
   REGION OUTPUTS
     // Write outputs
     IF (#statDisablingCompleted = TRUE) THEN
       // Reset outputs if disabling completed
       #statValid := FALSE;
       #statBusy := FALSE;
       #statError := FALSE;
       #statErrorUserCleared := FALSE;
       #statErrorAutoCleared := FALSE;
       #statStatus := #STATUS_NO_CALL;
       // TODO: Reset application specific outputs
       #statWaitMain := FALSE;

     ELSIF (#statErrorUserCleared = TRUE) AND (#statError = FALSE) THEN
       // Error can only be cleared by user; rising edge at enable input is needed to continue 
       #statValid := FALSE;
       #statBusy := FALSE;
       #statError := TRUE;
       #statFBState := #FB_STATE_NO_PROCESSING; // Switch state machine to "no processing"

     ELSIF (#statErrorAutoCleared = TRUE) AND (#statError = FALSE) THEN
       // Error can be reset by FB automatically  
       #statValid := FALSE;
       #statBusy := TRUE;
       #statError := TRUE;
       // TODO: Handling of autocleared error

     ELSIF (#statErrorAutoCleared = FALSE) AND (#statErrorUserCleared = FALSE) AND (#statError = TRUE) THEN
       // If autocleared error is acknowledged
       #statValid := TRUE;
       #statBusy := TRUE;
       #statError := FALSE;
       #statStatus := #STATUS_SUBSEQUENT_CALL;
     END_IF;

     // Write static values to outputs
     #valid := #statValid;
     #busy := #statBusy;
     #error := #statError;
     #status := #statStatus;
     // TODO: Write application specific static values to outputs
     #waitMain := #statWaitMain;
   END_REGION OUTPUTS
END_FUNCTION_BLOCK

FUNCTION "LKinCtrl_CheckPathDataCmd" : Word   // FC35000, SCL
TITLE = LKinCtrl_CheckPathDataCmd
{ S7_Optimized_Access := 'TRUE' }
AUTHOR : tech.team.motioncontrol@siemens.com
FAMILY : LKinCtrl
VERSION : 1.3
// The FC checks a PathData command to be configured correctly
   VAR_OUTPUT
      cmdIsMotionCmd : Bool;   // TRUE: Command is a motion command
   END_VAR
   VAR_IN_OUT
      pathDataCmd : Variant;   // variant for PathData command
   END_VAR
   VAR_TEMP
      tmpError : Bool;   // temporary variable for error bit
      tmpStatus : Word;   // temporary variable for status word
      tempFlagCtr : Int;   // temporary counter for flags
      tempPathDataCmd_regular : REF_TO "LKinCtrl_typePathDataElement";   // temporary reference to PathData element
      tempPathDataCmd_PreBuf : REF_TO "LKinCtrl_typePathDataElement_PreBuf";   // temporary reference to PathData_PreBuf element
      tempPathDataCmd_checking : "LKinCtrl_typePathDataElement";   // temporary variable for PathDataElement being checked
      tempPathDataType : Int;   // temporary variable storing detected PathData type
   END_VAR
   // Ret_Val : return value
   VAR CONSTANT
      STATUS_NO_ERROR_IN_COMMAND : Word := 16#0000;   // status no error found command
      ERR_PATHDATA_CMDTYPE : Word := 16#80A0;   // error due to wrong cmdType
      ERR_PATHDATA_COORDSYSTEM : Word := 16#80B1;   // error due to wrong coordinate system
      ERR_PATHDATA_VELOCITY : Word := 16#8003;   // error due to wrong velocity
      ERR_PATHDATA_ACCELERATION : Word := 16#8004;   // error due to wrong acceleration
      ERR_PATHDATA_DECELERATION : Word := 16#8005;   // error due to wrong deceleration
      ERR_PATHDATA_JERK : Word := 16#8006;   // error due to wrong jerk
      ERR_PATHDATA_ORIENTATIONDIRECTION : Word := 16#8007;   // error due to wrong orientation direction
      ERR_PATHDATA_BUFFERMODE : Word := 16#80B2;   // error due to wrong buffer mode
      ERR_PATHDATA_DYNAMICADAPTION : Word := 16#80B5;   // error due to wrong dynamic adaption
      ERR_PATHDATA_CIRCMODE : Word := 16#80B6;   // error due to wrong circle mode
      ERR_PATHDATA_PATHCHOICE : Word := 16#80B9;   // error due to wrong path choice
      ERR_PATHDATA_CIRCLEPLANE : Word := 16#80BA;   // error due to wrong circle plane
      ERR_PATHDATA_RADIUS : Word := 16#80BB;   // error due to wrong radius
      ERR_PATHDATA_ARC : Word := 16#80BC;   // error due to wrong arc
      ERR_PATHDATA_SETFLAGS_FLAG : Word := 16#80D1;   // error due to wrong set flag definition
      ERR_PATHDATA_SETFLAGS_FLAGMODE : Word := 16#80D2;   // error due to wrong set flag mode definition
      ERR_PATHDATA_VALUEFLAGS_FLAG : Word := 16#80D3;   // error due to wrong value flag definition
      ERR_PATHDATA_VALUEFLAGS_FLAGMODE : Word := 16#80D4;   // error due to wrong value flag mode definition
      ERR_PATHDATA_OFFSET_PARA_NO : Word := 16#80A1;   // error due to wrong offset parameter set number
      ERR_PATHDATA_OFFSET_MAINPATHPLANE : Word := 16#80A2;   // error due to wrong main path plane
      ERR_PATHDATA_POSITIONMODE : Word := 16#80A3;   // error due to wrong position mode
      ERR_PATHDATA_LINK_CONSTELLATION : Word := 16#80A4;   // error due to wrong link constellation
      ERR_PATHDATA_CONVEYOR_PARA_NO : Word := 16#80A5;   // error due to wrong conveyor parameter set number / error due to wrong link constellation
   END_VAR
BEGIN
   //==========================================================================================
   // SIEMENS AG
   // (c)Copyright 2020 All Rights Reserved
   //------------------------------------------------------------------------------------------
   // Library: LKinCtrl
   // Tested with: S7-1517T-3 PN/DP
   // Engineering: TIA Portal V15
   // Restrictions: ---
   // Requirements: S7-1500T FW 2.8
   // Functionality: LKinCtrl_CheckPathDataCmd
   // The FC checks a PathData command to be configured correctly
   // 
   // Support: tech.team.motioncontrol@siemens.com
   // Note: Parameter comments are only available in language 'English (United States)'
   //------------------------------------------------------------------------------------------
   // Change log table:
   // Version    Date          Expert in charge    Changes applied
   // 01.00.00   26.02.2019    JR                  First release version v1.0
   // 01.01.00   14.06.2019    JR                  added flagOnly command
   // 01.02.00   03.12.2019    JR                  added command checks for value flags
   // 01.02.01   30.01.2020    FR                  separate constant for flag arrays
   // 01.02.02   09.04.2020    FR                  copy valueFlags & CS to temp also
   // 01.03.00   16.04.2020    FR                  added moveDirect & trackConveyor
   //===========================================================================================

   // FC initialization
   //====================================================================================================================================
   #tmpError := FALSE;
   #tmpStatus := #STATUS_NO_ERROR_IN_COMMAND;

   // PathData conversion (reduced, regular(no suffix), advanced)
   //===========================================================================================
   REGION PATHDATA_ELEMENT_CONVERSION
     // regulat PathDataCommand
       IF TypeOf(#pathDataCmd) = LKinCtrl_typePathDataElement THEN
           // reference internal PathDataCommand to attached Variant
           #tempPathDataCmd_regular ?= #pathDataCmd;
           #tempPathDataType := 1;
           // copy to internal PathData (full version)
           #tempPathDataCmd_checking.cmdType := #tempPathDataCmd_regular<?OpDeref?>.cmdType;
           #tempPathDataCmd_checking.cmdCoordinates.coordSystem := #tempPathDataCmd_regular<?OpDeref?>.cmdCoordinates.coordSystem;
           #tempPathDataCmd_checking.cmdParameters := #tempPathDataCmd_regular<?OpDeref?>.cmdParameters;
           #tempPathDataCmd_checking.setFlags := #tempPathDataCmd_regular<?OpDeref?>.setFlags;
           #tempPathDataCmd_checking.valueFlags := #tempPathDataCmd_regular<?OpDeref?>.valueFlags;

           // PathDataPreBuffered PathDataCommand
       ELSIF TypeOf(#pathDataCmd) = LKinCtrl_typePathDataElement_PreBuf THEN
           #tempPathDataCmd_PreBuf ?= #pathDataCmd;
           #tempPathDataType := 2;
           // copy to internal PathData (full version)
           #tempPathDataCmd_checking.cmdType := #tempPathDataCmd_PreBuf<?OpDeref?>.cmdType;
           #tempPathDataCmd_checking.cmdCoordinates.coordSystem := #tempPathDataCmd_PreBuf<?OpDeref?>.cmdCoordinates.coordSystem;
           #tempPathDataCmd_checking.cmdParameters := #tempPathDataCmd_PreBuf<?OpDeref?>.cmdParameters;
           #tempPathDataCmd_checking.setFlags := #tempPathDataCmd_PreBuf<?OpDeref?>.setFlags;
           #tempPathDataCmd_checking.valueFlags := #tempPathDataCmd_PreBuf<?OpDeref?>.valueFlags;
       END_IF;
   END_REGION PATHDATA_CONVERSION 

   // PathData command 
   //====================================================================================================================================
   //PathData - command - cmdType
   // check for wrong PathData parameter cmdType
   IF (#tempPathDataCmd_checking.cmdType < "LKINCTRL_CMD_FLAG_ONLY"                      // lower limit MC cmdTypes
       OR #tempPathDataCmd_checking.cmdType > "LKINCTRL_MC_MOVEDIRECTREL")               // upper limit MC cmdTypes
     AND #tempPathDataCmd_checking.cmdType <> "LKINCTRL_CMD_WAIT_TIME"                   // exact cmdType constant for wait time
     AND #tempPathDataCmd_checking.cmdType <> "LKINCTRL_CONFIG_START_OFFSET_COMP_LEFT"   // exact cmdType constant for activation offset compensation left
     AND #tempPathDataCmd_checking.cmdType <> "LKINCTRL_CONFIG_START_OFFSET_COMP_RIGHT"  // exact cmdType constant for activation offset compensation right
     AND #tempPathDataCmd_checking.cmdType <> "LKINCTRL_CONFIG_END_OFFSET_COMP"          // exact cmdType constant for deactivation offset compensation
     AND #tempPathDataCmd_checking.cmdType <> "LKINCTRL_MC_TRACKCONVEYORBELT"
   THEN
     #tmpError := TRUE;
     #tmpStatus := #ERR_PATHDATA_CMDTYPE;
   END_IF;

   //PathData - command - cmdType
   // add separation for motion / non-motion commands here
   IF #tempPathDataCmd_checking.cmdType = "LKINCTRL_CMD_WAIT_TIME"
       OR #tempPathDataCmd_checking.cmdType = "LKINCTRL_CMD_FLAG_ONLY"
       OR #tempPathDataCmd_checking.cmdType = "LKINCTRL_MC_TRACKCONVEYORBELT"
     // add further non-motion commands here later (Zones, CS, ...)
     // only separate commands that will be copied to PathData_preBuffered
   THEN
     #cmdIsMotionCmd := FALSE;
   ELSE
     #cmdIsMotionCmd := TRUE;
   END_IF;

   //PathData - command - cmdCoordinates - coordSystem
   IF #tempPathDataCmd_checking.cmdType >= "LKINCTRL_MC_MOVELINEARABS"                           // lower limit path command cmdTypes
       AND #tempPathDataCmd_checking.cmdType <= "LKINCTRL_MC_MOVECIRCULARREL"                    // upper limit path command cmdTypes
   THEN
       // check for wrong parameter PathData coordSystem
       // CS is not WCS - OCS3 --> Error
       IF #tempPathDataCmd_checking.cmdCoordinates.coordSystem < "CS_WCS"
           OR #tempPathDataCmd_checking.cmdCoordinates.coordSystem > "CS_OCS3"
       THEN
           #tmpError := TRUE;
           #tmpStatus := #ERR_PATHDATA_COORDSYSTEM;
       END_IF;
   ELSIF #tempPathDataCmd_checking.cmdType >= "LKINCTRL_MC_MOVEDIRECTABS"                          // lower limit axis command cmdTypes
       AND #tempPathDataCmd_checking.cmdType <= "LKINCTRL_MC_MOVEDIRECTREL"                        // upper limit axis command cmdTypes
   THEN
       // check for wrong parameter PathData coordSystem
       // CS is not WCS - OCS3 and not MCS --> Error
       IF (#tempPathDataCmd_checking.cmdCoordinates.coordSystem < "CS_WCS"
           OR #tempPathDataCmd_checking.cmdCoordinates.coordSystem > "CS_OCS3")
           AND NOT (#tempPathDataCmd_checking.cmdCoordinates.coordSystem = "CS_MCS")
       THEN
           #tmpError := TRUE;
           #tmpStatus := #ERR_PATHDATA_COORDSYSTEM;
       END_IF;
       // Check conveyTracking coordinate system to be OCS1-3
   ELSIF #tempPathDataCmd_checking.cmdType = "LKINCTRL_MC_TRACKCONVEYORBELT"
       AND (#tempPathDataCmd_checking.cmdCoordinates.coordSystem < "CS_OCS1"
       OR #tempPathDataCmd_checking.cmdCoordinates.coordSystem > "CS_OCS3")
   THEN
       #tmpError := TRUE;
       #tmpStatus := #ERR_PATHDATA_COORDSYSTEM;
   END_IF;

   //PathData - command - cmdParameters - pathDynamics
   // Check MoveDirect dynamics
   IF #tempPathDataCmd_checking.cmdType >= "LKINCTRL_MC_MOVEDIRECTABS"                          // lower limit axis command cmdTypes
       AND #tempPathDataCmd_checking.cmdType <= "LKINCTRL_MC_MOVEDIRECTREL"                     // upper limit axis command cmdTypes
   THEN                
       // Check for wrong dynamics factors
       IF #tempPathDataCmd_checking.cmdParameters.pathDynamics.velocity > 1.0
           OR #tempPathDataCmd_checking.cmdParameters.pathDynamics.velocity = 0.0
       THEN
           #tmpError := TRUE;
           #tmpStatus := #ERR_PATHDATA_VELOCITY;
       END_IF;
       IF #tempPathDataCmd_checking.cmdParameters.pathDynamics.acceleration > 1.0
           OR #tempPathDataCmd_checking.cmdParameters.pathDynamics.acceleration = 0.0
       THEN
           #tmpError := TRUE;
           #tmpStatus := #ERR_PATHDATA_ACCELERATION;
       END_IF;
       IF #tempPathDataCmd_checking.cmdParameters.pathDynamics.deceleration > 1.0
           OR #tempPathDataCmd_checking.cmdParameters.pathDynamics.deceleration = 0.0
       THEN
           #tmpError := TRUE;
           #tmpStatus := #ERR_PATHDATA_DECELERATION;
       END_IF;
       IF (#tempPathDataCmd_checking.cmdParameters.pathDynamics.jerk > 0.0
           AND #tempPathDataCmd_checking.cmdParameters.pathDynamics.jerk < 0.1)
           OR #tempPathDataCmd_checking.cmdParameters.pathDynamics.jerk > 0.9
       THEN
           #tmpError := TRUE;
           #tmpStatus := #ERR_PATHDATA_JERK;
       END_IF;
   END_IF;

   //PathData - command - cmdParameters - orientationDirection
   // check for wrong parameter PathData orientationDirection
   IF #tempPathDataCmd_checking.cmdParameters.orientationDirection < 1
     OR #tempPathDataCmd_checking.cmdParameters.orientationDirection > 3
   THEN
     #tmpError := TRUE;
     #tmpStatus := #ERR_PATHDATA_ORIENTATIONDIRECTION;
   END_IF;

   //PathData - command - cmdParameters - bufferMode
   // check for wrong parameter PathData bufferMode
   IF #tempPathDataCmd_checking.cmdParameters.bufferMode <> 1
     AND #tempPathDataCmd_checking.cmdParameters.bufferMode <> 2
     AND #tempPathDataCmd_checking.cmdParameters.bufferMode <> 5
   THEN
     #tmpError := TRUE;
     #tmpStatus := #ERR_PATHDATA_BUFFERMODE;
   END_IF;

   //PathData - command - cmdParameters - dynamicAdaption
   // check for wrong parameter PathData dynamicAdaption
   IF #tempPathDataCmd_checking.cmdParameters.dynamicAdaption > 2
   THEN
     #tmpError := TRUE;
     #tmpStatus := #ERR_PATHDATA_DYNAMICADAPTION;
   END_IF;

   //PathData - command - circleParameter
   //====================================================================================================================================
   //PathData - command - circleParameter - circMode
   // check for wrong parameter PathData circMode
   IF #tempPathDataCmd_checking.cmdParameters.circleParameters.circMode < 0
     OR #tempPathDataCmd_checking.cmdParameters.circleParameters.circMode > 3
   THEN
     #tmpError := TRUE;
     #tmpStatus := #ERR_PATHDATA_CIRCMODE;
   END_IF;

   //PathData - command - circleParameter - pathChoice
   // check for wrong parameter PathData pathChoice
   IF #tempPathDataCmd_checking.cmdParameters.circleParameters.pathChoice < 0
     OR #tempPathDataCmd_checking.cmdParameters.circleParameters.pathChoice > 3
   THEN
     #tmpError := TRUE;
     #tmpStatus := #ERR_PATHDATA_PATHCHOICE;
   END_IF;

   //PathData - command - circleParameter - circlePlane
   // check for wrong parameter PathData circlePlane
   IF #tempPathDataCmd_checking.cmdParameters.circleParameters.circlePlane < 0
     OR #tempPathDataCmd_checking.cmdParameters.circleParameters.circlePlane > 2
   THEN
     #tmpError := TRUE;
     #tmpStatus := #ERR_PATHDATA_CIRCLEPLANE;
   END_IF;

   //PathData - command - circleParameter - radius
   // check for wrong parameter PathData radius
   IF #tempPathDataCmd_checking.cmdParameters.circleParameters.radius < 0.0
   THEN
     #tmpError := TRUE;
     #tmpStatus := #ERR_PATHDATA_RADIUS;
   END_IF;

   //PathData - command - circleParameter - arc
   // check for wrong parameter PathData arc
   IF #tempPathDataCmd_checking.cmdParameters.circleParameters.arc < 0.0
   THEN
     #tmpError := TRUE;
     #tmpStatus := #ERR_PATHDATA_ARC;
   END_IF;

   // PathData - command - moveDirect Parameters - linkConstellation
   IF #tempPathDataCmd_checking.cmdParameters.moveDirectParameters.linkConstellation <> 16#FFFF_FFFF
       AND #tempPathDataCmd_checking.cmdParameters.moveDirectParameters.linkConstellation > 16#0000_0007
   THEN
       #tmpError := TRUE;
       #tmpStatus := #ERR_PATHDATA_LINK_CONSTELLATION;
   END_IF;


   //PathData - command - moveDirect Parameters - positionMode
   IF #tempPathDataCmd_checking.cmdParameters.moveDirectParameters.positionMode < "PM_ABS_ABS"
       OR #tempPathDataCmd_checking.cmdParameters.moveDirectParameters.positionMode > "PM_ABS_REL"
   THEN
       #tmpError := TRUE;
       #tmpStatus := #ERR_PATHDATA_POSITIONMODE;
   END_IF;

   //PathData - command - offsetParameters - offSetParaNo
   // check for wrong parameter offSetParaNo
   IF (#tempPathDataCmd_checking.cmdType = "LKINCTRL_CONFIG_START_OFFSET_COMP_LEFT"
     OR #tempPathDataCmd_checking.cmdType = "LKINCTRL_CONFIG_START_OFFSET_COMP_RIGHT")
     AND (#tempPathDataCmd_checking.cmdParameters.offsetParameters.offsetParaNo < 1
     OR #tempPathDataCmd_checking.cmdParameters.offsetParameters.offsetParaNo > "LKINCTRL_NO_OF_OFFSETS")
   THEN
     #tmpError := TRUE;
     #tmpStatus := #ERR_PATHDATA_OFFSET_PARA_NO;
   END_IF;

   //PathData - command - offsetParameters - main
   // check for wrong parameter PathData circlePlane
   IF (#tempPathDataCmd_checking.cmdType = "LKINCTRL_CONFIG_START_OFFSET_COMP_LEFT"
     OR #tempPathDataCmd_checking.cmdType = "LKINCTRL_CONFIG_START_OFFSET_COMP_RIGHT")
     AND (#tempPathDataCmd_checking.cmdParameters.offsetParameters.mainPathPlane < 0
     OR #tempPathDataCmd_checking.cmdParameters.offsetParameters.mainPathPlane > 2)
   THEN
     #tmpError := TRUE;
     #tmpStatus := #ERR_PATHDATA_OFFSET_MAINPATHPLANE;
   END_IF;

   //PathData - command - conveyorParameters - conveyorParaNo
   IF #tempPathDataCmd_checking.cmdType = "LKINCTRL_MC_TRACKCONVEYORBELT"
       AND (#tempPathDataCmd_checking.cmdParameters.conveyorParameters.conveyorParaNo < 1
       OR #tempPathDataCmd_checking.cmdParameters.conveyorParameters.conveyorParaNo > "LKINCTRL_NO_OF_CONVEYOR")
   THEN
       #tmpError := TRUE;
       #tmpStatus := #ERR_PATHDATA_CONVEYOR_PARA_NO;
   END_IF;

   //PathData - command - setFlags
   //====================================================================================================================================
   FOR #tempFlagCtr := 1 TO "LKINCTRL_NO_OF_CMD_SETFLAGS" DO
     // check flag to be in range of flags InOut array at LKinCtrl_MC_MovePath
     IF #tempPathDataCmd_checking.setFlags[#tempFlagCtr].flag < -1
       OR #tempPathDataCmd_checking.setFlags[#tempFlagCtr].flag > "LKINCTRL_NO_OF_LAST_SETFLAG"
     THEN
       #tmpError := TRUE;
       #tmpStatus := #ERR_PATHDATA_SETFLAGS_FLAG;
       EXIT;
     END_IF;

     // check flagMode to be valid
     IF #tempPathDataCmd_checking.setFlags[#tempFlagCtr].flagMode <> 0
       AND #tempPathDataCmd_checking.setFlags[#tempFlagCtr].flagMode <> 1
       AND #tempPathDataCmd_checking.setFlags[#tempFlagCtr].flagMode <> 2
       AND #tempPathDataCmd_checking.setFlags[#tempFlagCtr].flagMode <> 3
       AND #tempPathDataCmd_checking.setFlags[#tempFlagCtr].flagMode <> 5
       AND #tempPathDataCmd_checking.setFlags[#tempFlagCtr].flagMode <> 10
       AND #tempPathDataCmd_checking.setFlags[#tempFlagCtr].flagMode <> 11
       AND #tempPathDataCmd_checking.setFlags[#tempFlagCtr].flagMode <> 13
       AND #tempPathDataCmd_checking.setFlags[#tempFlagCtr].flagMode <> 15
     THEN
       #tmpError := TRUE;
       #tmpStatus := #ERR_PATHDATA_SETFLAGS_FLAGMODE;
       EXIT;
     END_IF;
   END_FOR;

   //PathData - command - valueFlags
   //====================================================================================================================================
   FOR #tempFlagCtr := 1 TO "LKINCTRL_NO_OF_CMD_VALUEFLAGS" DO
     // check flag to be in range of flags InOut array at LKinCtrl_MC_MovePath
     IF #tempPathDataCmd_checking.valueFlags[#tempFlagCtr].flag < -1
       OR #tempPathDataCmd_checking.valueFlags[#tempFlagCtr].flag > "LKINCTRL_NO_OF_LAST_VALUEFLAG"
     THEN
       #tmpError := TRUE;
       #tmpStatus := #ERR_PATHDATA_VALUEFLAGS_FLAG;
       EXIT;
     END_IF;

     // check flagMode to be valid
     IF #tempPathDataCmd_checking.valueFlags[#tempFlagCtr].flagMode <> 0
       AND #tempPathDataCmd_checking.valueFlags[#tempFlagCtr].flagMode <> 1
       AND #tempPathDataCmd_checking.valueFlags[#tempFlagCtr].flagMode <> 2
       AND #tempPathDataCmd_checking.valueFlags[#tempFlagCtr].flagMode <> 3
       AND #tempPathDataCmd_checking.valueFlags[#tempFlagCtr].flagMode <> 5
       AND #tempPathDataCmd_checking.valueFlags[#tempFlagCtr].flagMode <> 10
       AND #tempPathDataCmd_checking.valueFlags[#tempFlagCtr].flagMode <> 11
       AND #tempPathDataCmd_checking.valueFlags[#tempFlagCtr].flagMode <> 13
       AND #tempPathDataCmd_checking.valueFlags[#tempFlagCtr].flagMode <> 15
     THEN
       #tmpError := TRUE;
       #tmpStatus := #ERR_PATHDATA_VALUEFLAGS_FLAGMODE;
       EXIT;
     END_IF;
   END_FOR;

   // Write Return Value
   //====================================================================================================================================
   IF #tmpError THEN
     #LKinCtrl_CheckPathDataCmd := #tmpStatus;
   ELSE
     #LKinCtrl_CheckPathDataCmd := #STATUS_NO_ERROR_IN_COMMAND;
   END_IF;
END_FUNCTION

FUNCTION "LKinCtrl_ConvElements_PathDataToPathData_PreBuf" : Void   // FC35002, SCL
TITLE = LKinCtrl_ConvElements_PathDataToPathData_PreBuf
{ S7_Optimized_Access := 'TRUE' }
AUTHOR : tech.team.motioncontrol@siemens.com
FAMILY : LKinCtrl
VERSION : 1.0
// The FC converts PathData commands to elements fitting the PathData_PreBuf structure
   VAR_INPUT
      copyCompensatedParametes : Bool;   // copy selection compensated parameters
      copyTransitionParameters : Bool;   // copy selection transition parameters
      copyFlags : Bool;   // copy selection flags
   END_VAR
   VAR_IN_OUT
      pathDataElement : "LKinCtrl_typePathDataElement";   // in: pathDataElement to be copied
      pathDataPreBufElement : "LKinCtrl_typePathDataElement_PreBuf";   // out: pathDataElement_PreBuf to be written
      pathDataName : String;   // name of PathData to be copied (separate from element)
   END_VAR
   VAR_TEMP
      tempFlagCtr : Int;
   END_VAR
BEGIN
   //==========================================================================================
   // SIEMENS AG
   // (c)Copyright 2019 All Rights Reserved
   //------------------------------------------------------------------------------------------
   // Library: LKinCtrl
   // Tested with: S7-1517T-3 PN/DP
   // Engineering: TIA Portal V15
   // Restrictions: ---
   // Requirements: S7-1500T FW 2.5
   // Functionality: LKinCtrl_ConvElements_PathDataToPathData_PreBuf
   // The FC converts PathData commands to elements fitting the PathData_PreBuf structure
   // 
   // Support: tech.team.motioncontrol@siemens.com
   // Note: Parameter comments are only available in language 'English (United States)'
   //------------------------------------------------------------------------------------------
   // Change log table:
   // Version    Date          Expert in charge    Changes applied
   // 01.00.00   20.02.2019    JR                  First release version v1.0
   // 01.00.01   16.08.2019    JR                  added setFlags edit code: flagMode: 3 -> 2
   // 01.00.02   28.01.2020    FR                  added value flags to copyFlags
   //===========================================================================================

   IF #copyCompensatedParametes THEN // copy target positions
     #pathDataPreBufElement.cmdCoordinates.absolutePosition[1] := #pathDataElement.cmdCoordinates.cartesianPosition.x;
     #pathDataPreBufElement.cmdCoordinates.absolutePosition[2] := #pathDataElement.cmdCoordinates.cartesianPosition.y;
     #pathDataPreBufElement.cmdCoordinates.absolutePosition[3] := #pathDataElement.cmdCoordinates.cartesianPosition.z;
     #pathDataPreBufElement.cmdCoordinates.absolutePosition[4] := #pathDataElement.cmdCoordinates.cartesianPosition.a;
     #pathDataPreBufElement.cmdCoordinates.coordSystem := #pathDataElement.cmdCoordinates.coordSystem;

     #pathDataPreBufElement.cmdParameters.circleParameters := #pathDataElement.cmdParameters.circleParameters;
   END_IF;


   #pathDataPreBufElement.cmdType := #pathDataElement.cmdType;
   #pathDataPreBufElement.cmdName := #pathDataElement.cmdName;
   #pathDataPreBufElement.pathDataName := #pathDataName;


   // copy equal command data type data
   #pathDataPreBufElement.cmdParameters.pathDynamics := #pathDataElement.cmdParameters.pathDynamics;
   #pathDataPreBufElement.cmdParameters.orientationDirection := #pathDataElement.cmdParameters.orientationDirection;
   #pathDataPreBufElement.cmdParameters.bufferMode := #pathDataElement.cmdParameters.bufferMode;
   IF #copyTransitionParameters THEN
     #pathDataPreBufElement.cmdParameters.transitionParameters := #pathDataElement.cmdParameters.transitionParameters;
   END_IF;

   #pathDataPreBufElement.cmdParameters.dynamicAdaption := #pathDataElement.cmdParameters.dynamicAdaption;

   IF #copyFlags THEN
     // Set flags (bool)
     // ---------------------------------------------------------------
     #pathDataPreBufElement.setFlags := #pathDataElement.setFlags;
     // // change flagMode 3 to flagMode 2 as functionality is equal
     // check for cmd to be flagOnly cmd
     // check for cmd to implement flag and flagMode to be flagMode 3
     FOR #tempFlagCtr := 1 TO "LKINCTRL_NO_OF_CMD_SETFLAGS" DO
       IF #pathDataPreBufElement.cmdType = "LKINCTRL_CMD_FLAG_ONLY"
         AND #pathDataPreBufElement.setFlags[#tempFlagCtr].flag <> -1
         AND #pathDataPreBufElement.setFlags[#tempFlagCtr].flagMode = 3
       THEN
         // change flagMode to flagMode 2
         #pathDataPreBufElement.setFlags[#tempFlagCtr].flagMode := 2;
       END_IF;
     END_FOR;
     // ---------------------------------------------------------------

     // Value flags (LReal)
     // ---------------------------------------------------------------
     #pathDataPreBufElement.valueFlags := #pathDataElement.valueFlags;
     // // change flagMode 3 to flagMode 2 as functionality is equal
     // check for cmd to be flagOnly cmd
     // check for cmd to implement flag and flagMode to be flagMode 3
     FOR #tempFlagCtr := 1 TO "LKINCTRL_NO_OF_CMD_VALUEFLAGS" DO
       IF #pathDataPreBufElement.cmdType = "LKINCTRL_CMD_FLAG_ONLY"
         AND #pathDataPreBufElement.valueFlags[#tempFlagCtr].flag <> -1
         AND #pathDataPreBufElement.valueFlags[#tempFlagCtr].flagMode = 3
       THEN
         // change flagMode to flagMode 2
         #pathDataPreBufElement.valueFlags[#tempFlagCtr].flagMode := 2;
       END_IF;
     END_FOR;
     // ---------------------------------------------------------------

   END_IF;
END_FUNCTION

FUNCTION "LKinCtrl_CalcResultingPos" : Word   // FC35003, SCL
TITLE = LKinCtrl_CalcResultingLastPos
{ S7_Optimized_Access := 'TRUE' }
AUTHOR : tech.team.motioncontrol@siemens.com
FAMILY : LKinCtrl
VERSION : 2.1
// The FC calculates the resulting last position after a given command being executed starting from a given 'previous' last position
   VAR_INPUT
      cmdType : Int;   // command type
      cartesianPos : Variant;   // cartesian position
      circleParameters : "LKinCtrl_typeCircleParameters";   // circle parameters
   END_VAR
   VAR_OUTPUT
      errorMessage : String;   // error message
   END_VAR
   VAR_IN_OUT
      lastAuxPoint : Array[1..3] of LReal;   // resulting auxPoint
      lastPos : Array[1..4] of LReal;   // resulting last position
   END_VAR
   VAR_TEMP
      tempCircRadiusPt1 : LReal;   // temporary variable for calculation
      tempCircRadiusPt2 : LReal;   // temporary variable for calculation
      tempCircRadiusPt3 : LReal;   // temporary variable for calculation
      tempCircRadius : LReal;   // temporary variable for calculation
      tempCircleDirectionSign : Int;   // temporary variable for calculation
      tempCtr : Int;   // temporary counter
      tempAngleRadius : LReal;   // temporary variable for calculation
      tempArgAcos : LReal;   // temporary variable for calculation
      tempCircMode3Selected : Bool;   // temporary variable for selected circMode
      tempArc : LReal;   // temporary variable for arc
      tempCartesianPosArray : REF_TO Array[1..4] of LReal;   // reference to coordinates from pre buf element
      tempCartesianPosStruct : REF_TO "LKinCtrl_typeCartesianPosition";   // reference to coordinates from normal element
      tempCartesianPos : Array[1..4] of LReal;   // temporary array for input end point
   END_VAR
   // Ret_Val : return value
   VAR CONSTANT
      ERR_INVALID_CMDTYPE : Word := 16#8264;   // error due to invalid cmdType
      ERR_INVALID_CIRCLEPLANE : Word := 16#8265;   // error due to invalid circle plane
      STATUS_NO_ERROR : Word := 16#0;   // status no error occured
   END_VAR
BEGIN
   //==========================================================================================
   // SIEMENS AG
   // (c)Copyright 2020 All Rights Reserved
   //------------------------------------------------------------------------------------------
   // Library: LKinCtrl
   // Tested with: S7-1517T-3 PN/DP
   // Engineering: TIA Portal V16
   // Restrictions: ---
   // Requirements: S7-1500T FW 2.8
   // Functionality: LKinCtrl_CalcResultingPos
   // The FC calculates the resulting last position after a given command being executed
   // starting from a given 'previous' last position 
   // 
   // Support: tech.team.motioncontrol@siemens.com
   // Note: Parameter comments are only available in language 'English (United States)'
   //------------------------------------------------------------------------------------------
   // Change log table:
   // Version    Date          Expert in charge    Changes applied
   // 01.00.00   11.03.2019    JR                  First release version v1.0
   // 01.00.01   17.05.2019    JR                  formal code changes fitting to styleguide
   // 02.00.00   06.04.2020    FR                  Changed interface to fit PathDataPreBuf and normal element; Also updated the calculation
   // 02.01.00   16.04.2020    FR                  Added moveDirect
   //===========================================================================================

   // Caclulation of resulting position after command
   //====================================================================================================================================
   REGION CALC_AND_STORE_LASTPOS
     // initially set return value to no error
     #LKinCtrl_CalcResultingPos := #STATUS_NO_ERROR;

     IF TypeOf(#cartesianPos) = LKinCtrl_typeCartesianPosition THEN
         // Assignment
         #tempCartesianPosStruct ?= #cartesianPos;

         // Assign temp with values
         #tempCartesianPos[1] := #tempCartesianPosStruct<?OpDeref?>.x;
         #tempCartesianPos[2] := #tempCartesianPosStruct<?OpDeref?>.y;
         #tempCartesianPos[3] := #tempCartesianPosStruct<?OpDeref?>.z;
         #tempCartesianPos[4] := #tempCartesianPosStruct<?OpDeref?>.a;

     ELSIF TypeOfElements(#cartesianPos) = LReal AND IS_ARRAY(#cartesianPos) AND CountOfElements(#cartesianPos) = 4 THEN
         // Assignment
         #tempCartesianPosArray ?= #cartesianPos;

         // Assign temp with values
         #tempCartesianPos := #tempCartesianPosArray<?OpDeref?>;

     ELSE
         ; // Wrong input ?
     END_IF;

     // calculate and store last target position
     IF #cmdType = "LKINCTRL_MC_MOVELINEARABS" OR #cmdType = "LKINCTRL_MC_MOVEDIRECTABS" THEN
         REGION LIN_ABS
             // directly copy given tarted position
             #lastPos := #tempCartesianPos;
         END_REGION LIN_ABS

     ELSIF #cmdType = "LKINCTRL_MC_MOVELINEARREL" OR #cmdType = "LKINCTRL_MC_MOVEDIRECTREL" THEN
         REGION LIN_REL
             // calculate resulting targetPosition for linear relative command
             FOR #tempCtr := 1 TO 4 DO
                 #lastPos[#tempCtr] := #lastPos[#tempCtr] + #tempCartesianPos[#tempCtr];
             END_FOR;
         END_REGION LIN_REL

     ELSIF #cmdType = "LKINCTRL_MC_MOVECIRCULARABS" OR #cmdType = "LKINCTRL_MC_MOVECIRCULARREL" THEN
       REGION CIRCULAR
         // calculate resulting targetPosition for circular absolute command
         // separation of circModes
         // circMode CM: 0 & CM: 2 & CM: 3
         IF #circleParameters.circMode = "CM_BORDER"
           OR #circleParameters.circMode = "LKINCTRL_CIRCMODE_GCODE" // conversion in COff section or LKinCtrl_MC_ExecuteKinMotionCmd
         THEN
           REGION CM_0_3
             IF #cmdType = "LKINCTRL_MC_MOVECIRCULARREL" THEN
               // Calculate absoulte EndPoint
               FOR #tempCtr := 1 TO 4 DO
                 #lastPos[#tempCtr] := #lastPos[#tempCtr] + #tempCartesianPos[#tempCtr];
               END_FOR;
               // Calculate absoulte AuxPoint
               FOR #tempCtr := 1 TO 3 DO
                 #lastAuxPoint[#tempCtr] := #lastPos[#tempCtr] + #circleParameters.auxPoint[#tempCtr];
               END_FOR;
             ELSE
               // directly copy given endPoint as LastPos
               #lastPos := #tempCartesianPos;
               // directly copy given auxPoint
               #lastAuxPoint := #circleParameters.auxPoint;
             END_IF;
           END_REGION CM_0_3

           // circMode CM: 1
         ELSIF #circleParameters.circMode = "CM_CENTER" THEN
           REGION CM_1
             // ============================================================================
             IF #cmdType = "LKINCTRL_MC_MOVECIRCULARREL" THEN
               // run same calculation to MC_MOVECIRCULARABS, but convert (rel -> abs) auxPoint before
               FOR #tempCtr := 1 TO 3 DO
                 #lastAuxPoint[#tempCtr] := #lastPos[#tempCtr] + #circleParameters.auxPoint[#tempCtr];
               END_FOR;
             ELSE
               // directly copy given auxPoint
               #lastAuxPoint := #circleParameters.auxPoint;
             END_IF;
             // ==============================================================================

             // Copy orientation position
             #lastPos[4] := #tempCartesianPos[4];

             // Copy arc to temp
             #tempArc := #circleParameters.arc;

             // check for angles bigger than full circle (360 degrees)
             IF #tempArc > 360.0 THEN
               // check for angles being multiple of 360 degrees (system commands do run bigger circles)
               #tempArc := LREAL_TO_DINT(#tempArc) MOD 360;
             END_IF;

             // try catching complete circles without calculation
             IF #tempArc = 360.0 OR #tempArc = 0.0 THEN
               // keep old positions, do nothing
               ;
             ELSE
               // run regular calculation

               // calculate radius of circle around auxPoint - new 
               // Added CaseSelection // FR 2019/04/17
               CASE #circleParameters.circlePlane OF
                 0:  // 0: "CP_XZ" - circle plane XZ
                   #tempCircRadiusPt1 := (#lastPos[1] - #lastAuxPoint[1]) * (#lastPos[1] - #lastAuxPoint[1]);
                   #tempCircRadiusPt2 := 0.0;//((lastPos[2] - lastAuxPoint[2]) * (lastPos[2] - lastAuxPoint[2]);
                   #tempCircRadiusPt3 := (#lastPos[3] - #lastAuxPoint[3]) * (#lastPos[3] - #lastAuxPoint[3]);
                 1:  // 1: "CP_YZ" - circle plane YZ
                   #tempCircRadiusPt1 := 0.0;//((lastPos[1] - lastAuxPoint[1]) * (lastPos[1] - lastAuxPoint[1]);
                   #tempCircRadiusPt2 := (#lastPos[2] - #lastAuxPoint[2]) * (#lastPos[2] - #lastAuxPoint[2]);
                   #tempCircRadiusPt3 := (#lastPos[3] - #lastAuxPoint[3]) * (#lastPos[3] - #lastAuxPoint[3]);
                 2:  // 2: "CP_XY" - circle plane XY
                   #tempCircRadiusPt1 := (#lastPos[1] - #lastAuxPoint[1]) * (#lastPos[1] - #lastAuxPoint[1]);
                   #tempCircRadiusPt2 := (#lastPos[2] - #lastAuxPoint[2]) * (#lastPos[2] - #lastAuxPoint[2]);
                   #tempCircRadiusPt3 := 0.0;//(lastPos[3] - lastAuxPoint[3]) * (lastPos[3] - lastAuxPoint[3]);
                 ELSE  // Statement section ELSE
                   // wrong circle plane, error will be caught earlier when checking PathDataElement
                   #LKinCtrl_CalcResultingPos := #ERR_INVALID_CIRCLEPLANE;
                   #errorMessage := 'invalid circle plane';
               END_CASE;

               #tempCircRadius := SQRT_LREAL(#tempCircRadiusPt1 + #tempCircRadiusPt2 + #tempCircRadiusPt3);

               // check for circleDirection -> define sign for motion command parameter 'arc'
               // 0: PC_Positive - positive direction (CCW)
               IF #circleParameters.pathChoice = 0 THEN
                 #tempCircleDirectionSign := 1;
                 // 1: PC_Negative - negative direction (CW)
               ELSIF #circleParameters.pathChoice = 1 THEN
                 #tempCircleDirectionSign := -1;
               END_IF;

               // rotation of vector between auxPoint and LastPos to get target position depending on circlePlane - new
               IF #tempCircMode3Selected = FALSE THEN
                 // 0: "CP_XZ" - circle plane XZ
                 IF #circleParameters.circlePlane = 0 THEN
                   #tempCircleDirectionSign *= -1;

                   // check circle radius not to be zero (avoid FPE)
                   IF #tempCircRadius <> 0 THEN
                     // calculate argument for ACOS (angle in between of two vectors - radius and x axis)
                     #tempArgAcos := ((#lastPos[1] - #lastAuxPoint[1]) * 1) / (#tempCircRadius * SQRT_LREAL(1));
                     // calculate ACOS for angle between to vectors
                     #tempAngleRadius := ACOS_LREAL(#tempArgAcos) * 180.0 / "LKINCTRL_PI";

                     // Added FR 2019/04/17: Was missing ?
                     IF #lastAuxPoint[3] > #lastPos[3] THEN
                       // acos result changed to negative angle
                       #tempAngleRadius := #tempAngleRadius * -1;
                       // check circle center point to be below (y direction) start point ==> not effective right now
                     ELSIF #lastAuxPoint[3] < #lastPos[3] THEN
                       #tempAngleRadius := #tempAngleRadius;
                     END_IF;

                   ELSE
                     // do not calculate angle in case of error; output status Message for internal debugging
                     #errorMessage := '#tempCircRadius = 0; AuxPoint is LastPosition';
                   END_IF;

                   #lastPos[1] := #tempCircRadius * COS_LREAL((#tempArc * #tempCircleDirectionSign + #tempAngleRadius) * "LKINCTRL_PI" / 180.0)
                   + #lastAuxPoint[1];
                   #lastPos[3] := #tempCircRadius * SIN_LREAL((#tempArc * #tempCircleDirectionSign + #tempAngleRadius) * "LKINCTRL_PI" / 180.0)
                   + #lastAuxPoint[3];

                   // 1: "CP_YZ" - circle plane YZ
                 ELSIF #circleParameters.circlePlane = 1 THEN
                   // check circle radius not to be zero (avoid FPE)
                   IF #tempCircRadius <> 0 THEN
                     // calculate argument for ACOS (angle in between of two vectors - radius and x axis)
                     #tempArgAcos := ((#lastPos[2] - #lastAuxPoint[2]) * 1) / (#tempCircRadius * SQRT_LREAL(1));
                     // calculate ACOS for angle between to vectors
                     #tempAngleRadius := ACOS_LREAL(#tempArgAcos) * 180.0 / "LKINCTRL_PI";

                     // Added FR 2019/04/17: Was missing ?
                     IF #lastAuxPoint[3] > #lastPos[3] THEN
                       // acos result changed to negative angle
                       #tempAngleRadius := #tempAngleRadius * -1;
                       // check circle center point to be below (y direction) start point ==> not effective right now
                     ELSIF #lastAuxPoint[3] < #lastPos[3] THEN
                       #tempAngleRadius := #tempAngleRadius;
                     END_IF;

                   ELSE
                     // do not calculate angle in case of error; output status Message for internal debugging
                     #errorMessage := '#tempCircRadius = 0; AuxPoint is LastPosition';
                   END_IF;

                   #lastPos[2] := #tempCircRadius * COS_LREAL((#tempArc * #tempCircleDirectionSign + #tempAngleRadius) * "LKINCTRL_PI" / 180.0)
                   + #lastAuxPoint[2];
                   #lastPos[3] := #tempCircRadius * SIN_LREAL((#tempArc * #tempCircleDirectionSign + #tempAngleRadius) * "LKINCTRL_PI" / 180.0)
                   + #lastAuxPoint[3];

                   // 2: "CP_XY" - circle plane XY
                 ELSIF #circleParameters.circlePlane = 2 THEN
                   // check circle radius not to be zero (avoid FPE)
                   IF #tempCircRadius <> 0 THEN
                     // calculate argument for ACOS (angle in between of two vectors - radius and x axis)
                     #tempArgAcos := ((#lastPos[1] - #lastAuxPoint[1]) * 1) / (#tempCircRadius * SQRT_LREAL(1));
                     // calculate ACOS for angle between to vectors
                     #tempAngleRadius := ACOS_LREAL(#tempArgAcos) * 180.0 / "LKINCTRL_PI";

                     // check statLastPos and AuxPoint to be in line parallel to y axis (separation of pos / neg angles)
                     //IF #tempArgAcos = 0 THEN // Commented Not necessary? FR 2019/04/17
                     // check circle center point to be above (y direction) start point
                     IF #lastAuxPoint[2] > #lastPos[2] THEN
                       // acos result changed to negative angle
                       #tempAngleRadius := #tempAngleRadius * -1;
                       // check circle center point to be below (y direction) start point ==> not effective right now
                     ELSIF #lastAuxPoint[2] < #lastPos[2] THEN // Changed > to < // FR 2019/04/17
                       #tempAngleRadius := #tempAngleRadius;
                     END_IF;
                     //END_IF;
                     //
                   ELSE
                     // do not calculate angle in case of error; output status Message for internal debugging
                     #errorMessage := '#tempCircRadius = 0; AuxPoint is LastPosition';
                   END_IF;

                   #lastPos[1] := #tempCircRadius * COS_LREAL((#tempArc * #tempCircleDirectionSign + #tempAngleRadius) * "LKINCTRL_PI" / 180.0)
                   + #lastAuxPoint[1];
                   #lastPos[2] := #tempCircRadius * SIN_LREAL((#tempArc * #tempCircleDirectionSign + #tempAngleRadius) * "LKINCTRL_PI" / 180.0)
                   + #lastAuxPoint[2];
                 END_IF;
               END_IF;

             END_IF;
           END_REGION CM_1

           // Circle mode 2 ==> define circle with radius and end point
         ELSIF #circleParameters.circMode = "CM_RADIUS" THEN
           REGION CM_2 
             IF #cmdType = "LKINCTRL_MC_MOVECIRCULARREL" THEN
               // changes JR: 2019/04/29 - only selective #lastPos writing
               // only write parameters for used planes ==> exclude unused plane coordinates for relative commands
               IF #circleParameters.circlePlane = 0 THEN   // XZ plane
                 #lastPos[1] += #tempCartesianPos[1];
                 // exclude y coordinate
                 #lastPos[3] += #tempCartesianPos[3];
               ELSIF #circleParameters.circlePlane = 1 THEN   // YZ plane
                 // exclude x coordinate
                 #lastPos[2] += #tempCartesianPos[2];
                 #lastPos[3] += #tempCartesianPos[3];
               ELSIF #circleParameters.circlePlane = 2 THEN   // XY plane
                 #lastPos[1] += #tempCartesianPos[1];
                 #lastPos[2] += #tempCartesianPos[2];
                 // exclude z coordinate
               END_IF;
               // Always write orientation
               #lastPos[4] += #tempCartesianPos[4];

             ELSE
               // changes JR: 2019/04/29 - only selective #lastPos writing
               // only write parameters for used planes ==> exclude unused plane coordinates for relative commands
               IF #circleParameters.circlePlane = 0 THEN   // XZ plane
                 #lastPos[1] := #tempCartesianPos[1];
                 // exclude y coordinate
                 #lastPos[3] := #tempCartesianPos[3];
               ELSIF #circleParameters.circlePlane = 1 THEN   // YZ plane
                 // exclude x coordinate
                 #lastPos[2] := #tempCartesianPos[2];
                 #lastPos[3] := #tempCartesianPos[3];
               ELSIF #circleParameters.circlePlane = 2 THEN   // XY plane
                 #lastPos[1] := #tempCartesianPos[1];
                 #lastPos[2] := #tempCartesianPos[2];
                 // exclude z coordinate
               END_IF;
               // Always write orientation
               #lastPos[4] := #tempCartesianPos[4];

             END_IF;
           END_REGION CM_2
         END_IF;
       END_REGION CIRCULAR

     ELSE
       // wrong cmdType
       #LKinCtrl_CalcResultingPos := #ERR_INVALID_CMDTYPE;
       #errorMessage := 'invalid cmdType';
     END_IF;
   END_REGION CALC_AND_STORE_LASTPOS
END_FUNCTION

FUNCTION "LKinCtrl_CheckForCmdLengthZero" : Void   // FC35004, SCL
TITLE = LKinCtrl_CheckForCmdLengthZero
{ S7_Optimized_Access := 'TRUE' }
AUTHOR : tech.team.motioncontrol@siemens.com
FAMILY : LKinCtrl
VERSION : 2.0
// The FC checks a PathData commands to have the length zero
   VAR_INPUT
      lastPos : Array[1..4] of LReal;   // starting position of command
   END_VAR
   VAR_OUTPUT
      commandLengthIsZero : Bool;   // TRUE: resulting command length is zero
   END_VAR
   VAR_IN_OUT
      command : "LKinCtrl_typePathDataElement";   // command to be checked
   END_VAR
BEGIN
   //==========================================================================================
   // SIEMENS AG
   // (c)Copyright 2020 All Rights Reserved
   //------------------------------------------------------------------------------------------
   // Library: LKinCtrl
   // Tested with: S7-1517T-3 PN/DP
   // Engineering: TIA Portal V15
   // Restrictions: ---
   // Requirements: S7-1500T FW 2.5
   // Functionality: LKinCtrl_CheckForCmdLengthZero
   // The FC checks a PathData commands to have the length zero
   // 
   // Support: tech.team.motioncontrol@siemens.com
   // Note: Parameter comments are only available in language 'English (United States)'
   //------------------------------------------------------------------------------------------
   // Change log table:
   // Version    Date          Expert in charge    Changes applied
   // 01.00.00   11.03.2019    JR                  First release version v1.0
   // 01.00.01   28.01.2020    FR                  Added flagOnlyCmd 
   // 02.00.00   07.04.2020    FR                  Removed previous command and added lastPos instead
   //===========================================================================================

   //Check for command to have length zero
   //====================================================================================================================================
   // check for relative command with no distance information
   IF #command.cmdType = "LKINCTRL_MC_MOVELINEARREL"
     AND #command.cmdCoordinates.cartesianPosition.x = 0.0
     AND #command.cmdCoordinates.cartesianPosition.y = 0.0
     AND #command.cmdCoordinates.cartesianPosition.z = 0.0
     AND #command.cmdCoordinates.cartesianPosition.a = 0.0
   THEN
     // set output
     #commandLengthIsZero := TRUE;
   // check for two linear absolute commands to same target position
   ELSIF #command.cmdType = "LKINCTRL_MC_MOVELINEARABS"
     AND #command.cmdCoordinates.cartesianPosition.x = #lastPos[1]
     AND #command.cmdCoordinates.cartesianPosition.y = #lastPos[2]
     AND #command.cmdCoordinates.cartesianPosition.z = #lastPos[3]
     AND #command.cmdCoordinates.cartesianPosition.a = #lastPos[4]
   THEN
     // set output
     #commandLengthIsZero := TRUE;
     // linRel_0 ==> linAbs(prePrePos)

   // check for wait command
   ELSIF #command.cmdType = "LKINCTRL_CMD_WAIT_TIME" THEN
     // set output
     #commandLengthIsZero := TRUE;

   // Check for flag only cmd
   ELSIF #command.cmdType = "LKINCTRL_CMD_FLAG_ONLY" THEN
     // set output
     #commandLengthIsZero := TRUE;

   ELSE
     // set output
     #commandLengthIsZero := FALSE;
   END_IF;
END_FUNCTION

